(* Logix 5000 project; controller PLC_MCC1300_75F1 vendor 1 type 14 code 166 rev 32.11; software revision 32.04; part 80 of 83 *)
(* tags used below, declared in another part *)
   GP_OB_InitializeMain : GP_OB_Initialize;
   M302SpeedUp : MAC_SpeedUp;
   M307A_M3_DR : AXIS_CIP_DRIVE;
   M307A_M4_DR : AXIS_CIP_DRIVE;
   M307B_M1_DR : AXIS_CIP_DRIVE;
   M307C_M1_DR : AXIS_CIP_DRIVE;
   TMP_dDirection : DINT;
   TMP_dTarget : DINT;
   TMP_rAcc : REAL;
   TMP_rDec : REAL;
   TMP_rSpeed : REAL;
   Z300_Conveyor : UDT_StandConv[29];
   Z300_Conveyor_IN_MOTION : MAC_Conveyor_ZC_IN_MOTION[29];
   Z300_Conveyor_OUT_MOTION : MAC_Conveyor_ZC_OUT_MOTION[29];
(* MotionLogic, continued *)

   24: [XIC(Z300_Conveyor[14].OUTPUT_xDriveEnable.[0]) XIO(Z300_Conveyor_OUT_MOTION[14].DR_MSO_M[0].ER) MSO(M307A_M3_DR,Z300_Conveyor_OUT_MOTION[14].DR_MSO_M[0]) ,XIO(Z300_Conveyor_OUT_MOTION[14].DR_MSO_M[0].EN) OTU(Z300_Conveyor_OUT_MOTION[14].DR_MSO_M[0].ER) ,XIO(Z300_Conveyor[14].OUTPUT_xDriveEnable.[0]) OTU(Z300_Conveyor_OUT_MOTION[14].DR_MSO_M[0].EN) XIO(Z300_Conveyor_OUT_MOTION[14].DR_MSF_M[0].ER) MSF(M307A_M3_DR,Z300_Conveyor_OUT_MOTION[14].DR_MSF_M[0]) ,XIO(Z300_Conveyor_OUT_MOTION[14].DR_MSF_M[0].EN) OTU(Z300_Conveyor_OUT_MOTION[14].DR_MSF_M[0].ER) ];
   25: MUL(Z300_Conveyor[14].AUX_rgrAcc_m_s2[0],1000,TMP_rAcc)MUL(Z300_Conveyor[14].AUX_rgrDec_m_s2[0],1000,TMP_rDec)DIV(Z300_Conveyor[14].AUX_rgdRequestSpeed_mm_min[0],60,TMP_rSpeed);
   26: XIC(Z300_Conveyor[14].OS_xStartCount.0)OTU(Z300_Conveyor_IN_MOTION[14].DR_MAR_M[0].PC)OTU(Z300_Conveyor_IN_MOTION[14].DR_MRP_M[0].DN);
   27: [XIC(Z300_Conveyor[14].OUTPUT_xRun.0) MOV(0,TMP_dDirection) ,XIC(Z300_Conveyor[14].OUTPUT_xReverse.0) MOV(1,TMP_dDirection) ][XIO(Z300_Conveyor_IN_MOTION[14].DR_MAR_M[0].PC) ,XIO(Z300_Conveyor_IN_MOTION[14].DR_MRP_M[0].DN) ,XIO(Z300_Conveyor[14].OUTPUT_xPositioning.0) ]MAJ(M307A_M3_DR,Z300_Conveyor_OUT_MOTION[14].DR_MAJ_M[0],TMP_dDirection,TMP_rSpeed,Units per sec,TMP_rAcc,Units per sec2,TMP_rDec,Units per sec2,Trapezoidal,TMP_rAcc,TMP_rDec,Units per sec3,Enabled,Programmed,0,None);
   28: XIC(Z300_Conveyor[14].OS_xStartCount.0)MRP(M307A_M3_DR,Z300_Conveyor_OUT_MOTION[14].DR_MRP_M[0],Absolute,Actual,0);
   29: [XIC(Z300_Conveyor_IN_MOTION[14].DR_MRP_M[0].DN) XIC(Z300_Conveyor[14].OUTPUT_xPositioning.0) [XIC(Z300_Conveyor[14].tmON_PhFilter[0].DN) ,XIC(Z300_Conveyor_IN_MOTION[14].DR_MAR_M[0].EN) ] MAR(M307A_M3_DR,Z300_Conveyor_OUT_MOTION[14].DR_MAR_M[0],Negative_Edge,Disabled,0,0,1) ,XIO(Z300_Conveyor[14].OUTPUT_xPositioning.0) MDR(M307A_M3_DR,Z300_Conveyor_OUT_MOTION[14].DR_MDR_M[0],1) ];
   30: XIC(Z300_Conveyor[14].OUTPUT_xPositioning.0)XIC(Z300_Conveyor_IN_MOTION[14].DR_MAR_M[0].PC)DIV(Z300_Conveyor[14].AUX_rgdTarget_cmm[0],100,TMP_dTarget)ADD(TMP_dTarget,M307A_M4_DR.Registration1Position,TMP_dTarget)MAM(M307A_M3_DR,Z300_Conveyor_OUT_MOTION[14].DR_MAM_M[0],0,TMP_dTarget,TMP_rSpeed,Units per sec,TMP_rAcc,Units per sec2,TMP_rDec,Units per sec2,Trapezoidal,TMP_rAcc,TMP_rDec,Units per sec3,Enabled,Programmed,0,None,0,0);
   31: [XIC(Z300_Conveyor[14].OUTPUT_xChangeSpeed.0) ,XIC(M302SpeedUp.OS_xChangeAccDec) ,XIC(GP_OB_InitializeMain.OUT_xOs_200ms) ][XIO(Z300_Conveyor[14].OUTPUT_xReverse.0) ,XIC(Z300_Conveyor[14].OUTPUT_xReverse.0) MUL(TMP_rSpeed,-1.0,TMP_rSpeed) ]MCD(M307A_M3_DR,Z300_Conveyor_OUT_MOTION[14].DR_MCD_M[0],Jog,Yes,TMP_rSpeed,Yes,TMP_rAcc,Yes,TMP_rDec,No,TMP_rAcc,No,TMP_rDec,Units per sec,Units per sec2,Units per sec2,Units per sec3);
   32: XIO(Z300_Conveyor[14].OUTPUT_xRun.0)XIO(Z300_Conveyor[14].OUTPUT_xReverse.0)[XIC(Z300_Conveyor_IN_MOTION[14].DR_MAJ_M[0].IP) MAS(M307A_M3_DR,Z300_Conveyor_OUT_MOTION[14].DR_MASjog_M[0],Jog,Yes,TMP_rDec,Units per sec2,No,TMP_rDec,Units per sec3) ,XIC(Z300_Conveyor_IN_MOTION[14].DR_MAM_M[0].IP) MAS(M307A_M3_DR,Z300_Conveyor_OUT_MOTION[14].DR_MASpos_M[0],Move,Yes,TMP_rDec,Units per sec2,No,TMP_rDec,Units per sec3) ,XIO(Z300_Conveyor_IN_MOTION[14].DR_MAJ_M[0].IP) XIO(Z300_Conveyor_IN_MOTION[14].DR_MAM_M[0].IP) XIO(Z300_Conveyor_IN_MOTION[14].DR_MASjog_M[0].IP) XIO(Z300_Conveyor_IN_MOTION[14].DR_MASpos_M[0].IP) MAS(M307A_M3_DR,Z300_Conveyor_OUT_MOTION[14].DR_MASall_M[0],All,Yes,TMP_rDec,Units per sec2,No,TMP_rDec,Units per sec3) ];
   // M307AM4
   33: NOP();
   34: XIC(Z300_Conveyor[15].OUTPUT_xDriveReset.0)MASR(M307A_M4_DR,Z300_Conveyor_OUT_MOTION[15].DR_MASR_M[0]);
   35: [XIC(Z300_Conveyor[15].OUTPUT_xDriveEnable.[0]) XIO(Z300_Conveyor_OUT_MOTION[15].DR_MSO_M[0].ER) MSO(M307A_M4_DR,Z300_Conveyor_OUT_MOTION[15].DR_MSO_M[0]) ,XIO(Z300_Conveyor_OUT_MOTION[15].DR_MSO_M[0].EN) OTU(Z300_Conveyor_OUT_MOTION[15].DR_MSO_M[0].ER) ,XIO(Z300_Conveyor[15].OUTPUT_xDriveEnable.[0]) OTU(Z300_Conveyor_OUT_MOTION[15].DR_MSO_M[0].EN) XIO(Z300_Conveyor_OUT_MOTION[15].DR_MSF_M[0].ER) MSF(M307A_M4_DR,Z300_Conveyor_OUT_MOTION[15].DR_MSF_M[0]) ,XIO(Z300_Conveyor_OUT_MOTION[15].DR_MSF_M[0].EN) OTU(Z300_Conveyor_OUT_MOTION[15].DR_MSF_M[0].ER) ];
   36: MUL(Z300_Conveyor[15].AUX_rgrAcc_m_s2[0],1000,TMP_rAcc)MUL(Z300_Conveyor[15].AUX_rgrDec_m_s2[0],1000,TMP_rDec)DIV(Z300_Conveyor[15].AUX_rgdRequestSpeed_mm_min[0],60,TMP_rSpeed);
   37: XIC(Z300_Conveyor[15].OS_xStartCount.0)OTU(Z300_Conveyor_IN_MOTION[15].DR_MAR_M[0].PC)OTU(Z300_Conveyor_IN_MOTION[15].DR_MRP_M[0].DN);
   38: [XIC(Z300_Conveyor[15].OUTPUT_xRun.0) MOV(0,TMP_dDirection) ,XIC(Z300_Conveyor[15].OUTPUT_xReverse.0) MOV(1,TMP_dDirection) ][XIO(Z300_Conveyor_IN_MOTION[15].DR_MAR_M[0].PC) ,XIO(Z300_Conveyor_IN_MOTION[15].DR_MRP_M[0].DN) ,XIO(Z300_Conveyor[15].OUTPUT_xPositioning.0) ]MAJ(M307A_M4_DR,Z300_Conveyor_OUT_MOTION[15].DR_MAJ_M[0],TMP_dDirection,TMP_rSpeed,Units per sec,TMP_rAcc,Units per sec2,TMP_rDec,Units per sec2,Trapezoidal,TMP_rAcc,TMP_rDec,Units per sec3,Enabled,Programmed,0,None);
   39: XIC(Z300_Conveyor[15].OS_xStartCount.0)MRP(M307A_M4_DR,Z300_Conveyor_OUT_MOTION[15].DR_MRP_M[0],Absolute,Actual,0);
   40: [XIC(Z300_Conveyor_IN_MOTION[15].DR_MRP_M[0].DN) XIC(Z300_Conveyor[15].OUTPUT_xPositioning.0) [XIC(Z300_Conveyor[15].tmON_PhFilter[0].DN) ,XIC(Z300_Conveyor_IN_MOTION[15].DR_MAR_M[0].EN) ] MAR(M307A_M4_DR,Z300_Conveyor_OUT_MOTION[15].DR_MAR_M[0],Negative_Edge,Disabled,0,0,1) ,XIO(Z300_Conveyor[14].OUTPUT_xPositioning.0) MDR(M307A_M4_DR,Z300_Conveyor_OUT_MOTION[15].DR_MDR_M[0],1) ];
   41: XIC(Z300_Conveyor[15].OUTPUT_xPositioning.0)XIC(Z300_Conveyor_IN_MOTION[15].DR_MAR_M[0].PC)DIV(Z300_Conveyor[15].AUX_rgdTarget_cmm[0],100,TMP_dTarget)ADD(TMP_dTarget,M307A_M4_DR.Registration1Position,TMP_dTarget)MAM(M307A_M4_DR,Z300_Conveyor_OUT_MOTION[15].DR_MAM_M[0],0,TMP_dTarget,TMP_rSpeed,Units per sec,TMP_rAcc,Units per sec2,TMP_rDec,Units per sec2,Trapezoidal,TMP_rAcc,TMP_rDec,Units per sec3,Enabled,Programmed,0,None,0,0);
   42: [XIC(Z300_Conveyor[15].OUTPUT_xChangeSpeed.0) ,XIC(M302SpeedUp.OS_xChangeAccDec) ,XIC(GP_OB_InitializeMain.OUT_xOs_200ms) ][XIO(Z300_Conveyor[15].OUTPUT_xReverse.0) ,XIC(Z300_Conveyor[15].OUTPUT_xReverse.0) MUL(TMP_rSpeed,-1.0,TMP_rSpeed) ]MCD(M307A_M4_DR,Z300_Conveyor_OUT_MOTION[15].DR_MCD_M[0],Jog,Yes,TMP_rSpeed,Yes,TMP_rAcc,Yes,TMP_rDec,No,TMP_rAcc,No,TMP_rDec,Units per sec,Units per sec2,Units per sec2,Units per sec3);
   43: XIO(Z300_Conveyor[15].OUTPUT_xRun.0)XIO(Z300_Conveyor[15].OUTPUT_xReverse.0)[XIC(Z300_Conveyor_IN_MOTION[15].DR_MAJ_M[0].IP) MAS(M307A_M4_DR,Z300_Conveyor_OUT_MOTION[15].DR_MASjog_M[0],Jog,Yes,TMP_rDec,Units per sec2,No,TMP_rDec,Units per sec3) ,XIC(Z300_Conveyor_IN_MOTION[15].DR_MAM_M[0].IP) MAS(M307A_M4_DR,Z300_Conveyor_OUT_MOTION[15].DR_MASpos_M[0],Move,Yes,TMP_rDec,Units per sec2,No,TMP_rDec,Units per sec3) ,XIO(Z300_Conveyor_IN_MOTION[15].DR_MAJ_M[0].IP) XIO(Z300_Conveyor_IN_MOTION[15].DR_MAM_M[0].IP) XIO(Z300_Conveyor_IN_MOTION[15].DR_MASjog_M[0].IP) XIO(Z300_Conveyor_IN_MOTION[15].DR_MASpos_M[0].IP) MAS(M307A_M4_DR,Z300_Conveyor_OUT_MOTION[15].DR_MASall_M[0],All,Yes,TMP_rDec,Units per sec2,No,TMP_rDec,Units per sec3) ];
END_ROUTINE

ROUTINE M307B_Motion   (* ladder *)
   // M307BM1
   0: NOP();
   1: XIC(Z300_Conveyor[16].OUTPUT_xDriveReset.0)MASR(M307B_M1_DR,Z300_Conveyor_OUT_MOTION[16].DR_MASR_M[0]);
   2: [XIC(Z300_Conveyor[16].OUTPUT_xDriveEnable.[0]) XIO(Z300_Conveyor_OUT_MOTION[16].DR_MSO_M[0].ER) MSO(M307B_M1_DR,Z300_Conveyor_OUT_MOTION[16].DR_MSO_M[0]) ,XIO(Z300_Conveyor_OUT_MOTION[16].DR_MSO_M[0].EN) OTU(Z300_Conveyor_OUT_MOTION[16].DR_MSO_M[0].ER) ,XIO(Z300_Conveyor[16].OUTPUT_xDriveEnable.[0]) OTU(Z300_Conveyor_OUT_MOTION[16].DR_MSO_M[0].EN) XIO(Z300_Conveyor_OUT_MOTION[16].DR_MSF_M[0].ER) MSF(M307B_M1_DR,Z300_Conveyor_OUT_MOTION[16].DR_MSF_M[0]) ,XIO(Z300_Conveyor_OUT_MOTION[16].DR_MSF_M[0].EN) OTU(Z300_Conveyor_OUT_MOTION[16].DR_MSF_M[0].ER) ];
   3: MUL(Z300_Conveyor[16].AUX_rgrAcc_m_s2[0],1000,TMP_rAcc)MUL(Z300_Conveyor[16].AUX_rgrDec_m_s2[0],1000,TMP_rDec)DIV(Z300_Conveyor[16].AUX_rgdRequestSpeed_mm_min[0],60,TMP_rSpeed);
   4: XIC(Z300_Conveyor[16].OS_xStartCount.0)OTU(Z300_Conveyor_IN_MOTION[16].DR_MAR_M[0].PC)OTU(Z300_Conveyor_IN_MOTION[16].DR_MRP_M[0].DN);
   5: [XIC(Z300_Conveyor[16].OUTPUT_xRun.0) MOV(0,TMP_dDirection) ,XIC(Z300_Conveyor[16].OUTPUT_xReverse.0) MOV(1,TMP_dDirection) ][XIO(Z300_Conveyor_IN_MOTION[16].DR_MAR_M[0].PC) ,XIO(Z300_Conveyor_IN_MOTION[16].DR_MRP_M[0].DN) ,XIO(Z300_Conveyor[16].OUTPUT_xPositioning.0) ]MAJ(M307B_M1_DR,Z300_Conveyor_OUT_MOTION[16].DR_MAJ_M[0],TMP_dDirection,TMP_rSpeed,Units per sec,TMP_rAcc,Units per sec2,TMP_rDec,Units per sec2,Trapezoidal,TMP_rAcc,TMP_rDec,Units per sec3,Enabled,Programmed,0,None);
   6: XIC(Z300_Conveyor[16].OS_xStartCount.0)MRP(M307B_M1_DR,Z300_Conveyor_OUT_MOTION[16].DR_MRP_M[0],Absolute,Actual,0);
   7: [XIC(Z300_Conveyor_IN_MOTION[16].DR_MRP_M[0].DN) XIC(Z300_Conveyor[16].OUTPUT_xPositioning.0) [XIC(Z300_Conveyor[16].tmON_PhFilter[0].DN) ,XIC(Z300_Conveyor_IN_MOTION[16].DR_MAR_M[0].EN) ] MAR(M307B_M1_DR,Z300_Conveyor_OUT_MOTION[16].DR_MAR_M[0],Negative_Edge,Disabled,0,0,1) ,XIO(Z300_Conveyor[16].OUTPUT_xPositioning.0) MDR(M307B_M1_DR,Z300_Conveyor_OUT_MOTION[16].DR_MDR_M[0],1) ];
   8: XIC(Z300_Conveyor[16].OUTPUT_xPositioning.0)XIC(Z300_Conveyor_IN_MOTION[16].DR_MAR_M[0].PC)DIV(Z300_Conveyor[16].AUX_rgdTarget_cmm[0],100,TMP_dTarget)ADD(TMP_dTarget,M307B_M1_DR.Registration1Position,TMP_dTarget)MAM(M307B_M1_DR,Z300_Conveyor_OUT_MOTION[16].DR_MAM_M[0],0,TMP_dTarget,TMP_rSpeed,Units per sec,TMP_rAcc,Units per sec2,TMP_rDec,Units per sec2,Trapezoidal,TMP_rAcc,TMP_rDec,Units per sec3,Enabled,Programmed,0,None,0,0);
   9: [XIC(Z300_Conveyor[16].OUTPUT_xChangeSpeed.0) ,XIC(M302SpeedUp.OS_xChangeAccDec) ,XIC(GP_OB_InitializeMain.OUT_xOs_200ms) ][XIO(Z300_Conveyor[16].OUTPUT_xReverse.0) ,XIC(Z300_Conveyor[16].OUTPUT_xReverse.0) MUL(TMP_rSpeed,-1.0,TMP_rSpeed) ]MCD(M307B_M1_DR,Z300_Conveyor_OUT_MOTION[16].DR_MCD_M[0],Jog,Yes,TMP_rSpeed,Yes,TMP_rAcc,Yes,TMP_rDec,No,TMP_rAcc,No,TMP_rDec,Units per sec,Units per sec2,Units per sec2,Units per sec3);
   10: XIO(Z300_Conveyor[16].OUTPUT_xRun.0)XIO(Z300_Conveyor[16].OUTPUT_xReverse.0)[XIC(Z300_Conveyor_IN_MOTION[16].DR_MAJ_M[0].IP) MAS(M307B_M1_DR,Z300_Conveyor_OUT_MOTION[16].DR_MASjog_M[0],Jog,Yes,TMP_rDec,Units per sec2,No,TMP_rDec,Units per sec3) ,XIC(Z300_Conveyor_IN_MOTION[16].DR_MAM_M[0].IP) MAS(M307B_M1_DR,Z300_Conveyor_OUT_MOTION[16].DR_MASpos_M[0],Move,Yes,TMP_rDec,Units per sec2,No,TMP_rDec,Units per sec3) ,XIO(Z300_Conveyor_IN_MOTION[16].DR_MAJ_M[0].IP) XIO(Z300_Conveyor_IN_MOTION[16].DR_MAM_M[0].IP) XIO(Z300_Conveyor_IN_MOTION[16].DR_MASjog_M[0].IP) XIO(Z300_Conveyor_IN_MOTION[16].DR_MASpos_M[0].IP) MAS(M307B_M1_DR,Z300_Conveyor_OUT_MOTION[16].DR_MASall_M[0],All,Yes,TMP_rDec,Units per sec2,No,TMP_rDec,Units per sec3) ];
END_ROUTINE

ROUTINE M307C_Motion   (* ladder *)
   // M307CM1
   0: NOP();
   1: XIC(Z300_Conveyor[17].OUTPUT_xDriveReset.0)MASR(M307C_M1_DR,Z300_Conveyor_OUT_MOTION[17].DR_MASR_M[0]);
   2: [XIC(Z300_Conveyor[17].OUTPUT_xDriveEnable.[0]) XIO(Z300_Conveyor_OUT_MOTION[17].DR_MSO_M[0].ER) MSO(M307C_M1_DR,Z300_Conveyor_OUT_MOTION[17].DR_MSO_M[0]) ,XIO(Z300_Conveyor_OUT_MOTION[17].DR_MSO_M[0].EN) OTU(Z300_Conveyor_OUT_MOTION[17].DR_MSO_M[0].ER) ,XIO(Z300_Conveyor[17].OUTPUT_xDriveEnable.[0]) OTU(Z300_Conveyor_OUT_MOTION[17].DR_MSO_M[0].EN) XIO(Z300_Conveyor_OUT_MOTION[17].DR_MSF_M[0].ER) MSF(M307C_M1_DR,Z300_Conveyor_OUT_MOTION[17].DR_MSF_M[0]) ,XIO(Z300_Conveyor_OUT_MOTION[17].DR_MSF_M[0].EN) OTU(Z300_Conveyor_OUT_MOTION[17].DR_MSF_M[0].ER) ];
   3: MUL(Z300_Conveyor[17].AUX_rgrAcc_m_s2[0],1000,TMP_rAcc)MUL(Z300_Conveyor[17].AUX_rgrDec_m_s2[0],1000,TMP_rDec)DIV(Z300_Conveyor[17].AUX_rgdRequestSpeed_mm_min[0],60,TMP_rSpeed);
   4: XIC(Z300_Conveyor[17].OS_xStartCount.0)OTU(Z300_Conveyor_IN_MOTION[17].DR_MAR_M[0].PC)OTU(Z300_Conveyor_IN_MOTION[17].DR_MRP_M[0].DN);
   5: [XIC(Z300_Conveyor[17].OUTPUT_xRun.0) MOV(0,TMP_dDirection) ,XIC(Z300_Conveyor[17].OUTPUT_xReverse.0) MOV(1,TMP_dDirection) ][XIO(Z300_Conveyor_IN_MOTION[17].DR_MAR_M[0].PC) ,XIO(Z300_Conveyor_IN_MOTION[17].DR_MRP_M[0].DN) ,XIO(Z300_Conveyor[17].OUTPUT_xPositioning.0) ]MAJ(M307C_M1_DR,Z300_Conveyor_OUT_MOTION[17].DR_MAJ_M[0],TMP_dDirection,TMP_rSpeed,Units per sec,TMP_rAcc,Units per sec2,TMP_rDec,Units per sec2,Trapezoidal,TMP_rAcc,TMP_rDec,Units per sec3,Enabled,Programmed,0,None);
   6: XIC(Z300_Conveyor[17].OS_xStartCount.0)MRP(M307C_M1_DR,Z300_Conveyor_OUT_MOTION[17].DR_MRP_M[0],Absolute,Actual,0);
   7: [XIC(Z300_Conveyor_IN_MOTION[17].DR_MRP_M[0].DN) XIC(Z300_Conveyor[17].OUTPUT_xPositioning.0) [XIC(Z300_Conveyor[17].tmON_PhFilter[0].DN) ,XIC(Z300_Conveyor_IN_MOTION[17].DR_MAR_M[0].EN) ] MAR(M307C_M1_DR,Z300_Conveyor_OUT_MOTION[17].DR_MAR_M[0],Negative_Edge,Disabled,0,0,1) ,XIO(Z300_Conveyor[17].OUTPUT_xPositioning.0) MDR(M307C_M1_DR,Z300_Conveyor_OUT_MOTION[17].DR_MDR_M[0],1) ];
   8: XIC(Z300_Conveyor[17].OUTPUT_xPositioning.0)XIC(Z300_Conveyor_IN_MOTION[17].DR_MAR_M[0].PC)DIV(Z300_Conveyor[17].AUX_rgdTarget_cmm[0],100,TMP_dTarget)ADD(TMP_dTarget,M307C_M1_DR.Registration1Position,TMP_dTarget)MAM(M307C_M1_DR,Z300_Conveyor_OUT_MOTION[17].DR_MAM_M[0],0,TMP_dTarget,TMP_rSpeed,Units per sec,TMP_rAcc,Units per sec2,TMP_rDec,Units per sec2,Trapezoidal,TMP_rAcc,TMP_rDec,Units per sec3,Enabled,Programmed,0,None,0,0);
   9: [XIC(Z300_Conveyor[17].OUTPUT_xChangeSpeed.0) ,XIC(M302SpeedUp.OS_xChangeAccDec) ,XIC(GP_OB_InitializeMain.OUT_xOs_200ms) ][XIO(Z300_Conveyor[17].OUTPUT_xReverse.0) ,XIC(Z300_Conveyor[17].OUTPUT_xReverse.0) MUL(TMP_rSpeed,-1.0,TMP_rSpeed) ]MCD(M307C_M1_DR,Z300_Conveyor_OUT_MOTION[17].DR_MCD_M[0],Jog,Yes,TMP_rSpeed,Yes,TMP_rAcc,Yes,TMP_rDec,No,TMP_rAcc,No,TMP_rDec,Units per sec,Units per sec2,Units per sec2,Units per sec3);
   10: XIO(Z300_Conveyor[17].OUTPUT_xRun.0)XIO(Z300_Conveyor[17].OUTPUT_xReverse.0)[XIC(Z300_Conveyor_IN_MOTION[17].DR_MAJ_M[0].IP) MAS(M307C_M1_DR,Z300_Conveyor_OUT_MOTION[17].DR_MASjog_M[0],Jog,Yes,TMP_rDec,Units per sec2,No,TMP_rDec,Units per sec3) ,XIC(Z300_Conveyor_IN_MOTION[17].DR_MAM_M[0].IP) MAS(M307C_M1_DR,Z300_Conveyor_OUT_MOTION[17].DR_MASpos_M[0],Move,Yes,TMP_rDec,Units per sec2,No,TMP_rDec,Units per sec3) ,XIO(Z300_Conveyor_IN_MOTION[17].DR_MAJ_M[0].IP) XIO(Z300_Conveyor_IN_MOTION[17].DR_MAM_M[0].IP) XIO(Z300_Conveyor_IN_MOTION[17].DR_MASjog_M[0].IP) XIO(Z300_Conveyor_IN_MOTION[17].DR_MASpos_M[0].IP) MAS(M307C_M1_DR,Z300_Conveyor_OUT_MOTION[17].DR_MASall_M[0],All,Yes,TMP_rDec,Units per sec2,No,TMP_rDec,Units per sec3) ];
END_ROUTINE
